VERSION : 0.1
// Data area for auto sequence timers
   VAR
      CV341_CLSD_DLY : TON_TIME;   // For the delay prior to the BC start command
      P305_STRTD_DLY : TON_TIME;   // For the delay after P305 has started
      P304_STRTD_DLY : TON_TIME;   // For the delay after P304 has started
      P303_STRTD_DLY : TON_TIME;   // For the delay after P304 has started
      PRE_GCU_TNK_FILL_DLY : TON_TIME;   // For the delay prior to GCU tank fill timer
      GCU_TNK_MAX_FILL_TMR : TON_TIME;   // For the maximum GCU fill time
      P305_STPD_DLY : TON_TIME;   // For the delay after P305 has stopped
      P304_STPD_DLY : TON_TIME;   // For the delay after P304 has stopped
      CV358_CLSD_DLY : TON_TIME;   // For the delay prior to the BC start command
      E400_STRTD_DLY : TON_TIME;   // For the delay after E400 has started
      E400_RNG_DLY : TON_TIME;   // For the delay as E400 runs at load
      CV401_OPND_DLY : TON_TIME;   // For the delay after CV401 has opened
      CV401_CLSD_DLY : TON_TIME;   // For the delay after CV401 has closed
      CV441_OPND_DLY : TON_TIME;   // For the delay after CV441 has opened
      CV441_CLSD_DLY : TON_TIME;   // For the delay after CV441 has closed
      PRE_441_OPN_DLY : TON_TIME;   // For the delay prior to CV441 opening
      VLV_CNFG_DN_DLY : TON_TIME;   // For the delay once the DeOx/ReOx are done
      CV405_OPND_DLY : TON_TIME;   // For the delay after CV405 has opened
      CV406_CLSD_DLY : TON_TIME;   // For the delay after CV406 has closed
      E400_STOP_TMR : TON_TIME;   // For the maximum PGC stop time
      P303_STPD_DLY : TON_TIME;   // For the maximum P303 stop time
      CV341_OPND_DLY : TON_TIME;   // For the delay after CV341 has opened
      GCU_TNK_MAX_DRN_TMR : TON_TIME;   // For the maximum GCU drain time
      POST_FLUSH_DLY : TON_TIME;   // Dor the delay after the tank has flushed
      "LIT304 Delay" : TON_TIME;
      P301_START_DLY : TON_TIME;   // Delay after starting the CSW pump
      "FS332 Delay" : TON_TIME;
      "Pre-Dwel PPPuls" : TP_TIME;
      SFTY_SYS_IL : TOF_TIME;
      OVR_TANK : TON_TIME;
      "Tank Close Delay" : TON_TIME;
   END_VAR
BEGIN
   CV341_CLSD_DLY.PT := T#10s;
   P305_STRTD_DLY.PT := T#5s;
   P304_STRTD_DLY.PT := T#5s;
   PRE_GCU_TNK_FILL_DLY.PT := T#15s;
   GCU_TNK_MAX_FILL_TMR.PT := T#300s;
   P305_STPD_DLY.PT := T#5s;
   P304_STPD_DLY.PT := T#5s;
   CV358_CLSD_DLY.PT := T#5s;
   P303_STRTD_DLY.PT := T#15s;
   E400_STRTD_DLY.PT := T#15s;
   E400_RNG_DLY.PT := T#5s;
   VLV_CNFG_DN_DLY.PT := T#10s;
   PRE_441_OPN_DLY.PT := T#15s;
   CV441_CLSD_DLY.PT := T#5s;
   CV441_OPND_DLY.PT := T#5s;
   CV401_CLSD_DLY.PT := T#5s;
   CV401_OPND_DLY.PT := T#5s;
   CV405_OPND_DLY.PT := T#10s;
   CV406_CLSD_DLY.PT := T#2s;
   E400_STOP_TMR.PT := T#180s;
   P303_STPD_DLY.PT := T#30s;
   CV341_OPND_DLY.PT := T#2s;
   GCU_TNK_MAX_DRN_TMR.PT := T#180s;
   POST_FLUSH_DLY.PT := T#60s;
   OVR_TANK.PT := T#1s;
   "Tank Close Delay".PT := T#1s;
END_DATA_BLOCK

// folder: 50 - 59 PLC Communication

DATA_BLOCK "51_SLAVE_STATUS"   // DB51
TITLE = Slave Status Data
{ S7_Optimized_Access := 'FALSE' }
AUTHOR : JRS
VERSION : 0.1
// Data area for status from slave PLC
   VAR
      HEART_BEAT : Bool;
      AUT_SEQ_RNG : Bool;   // Auto sequence running
      CRNT_MODE : Int := 1;   // 1 = Auto, 2 = Man, 3 = FatAuto, 4 = FatMan
      STARTING : Bool;   // IGG Is starting
      O2_LVL_OK : Bool;   // O2 Level within specification
      RUNNING : Bool;   // Running
      VLVS_AT_INIT : Bool;   // 1 = Valves at initial, 0 = Not
      ESTOP_OK : Bool;   // 1 = OK, 0 = Estop active
      IGG_ALARM : Bool;   // 1 = IGG Alarm state, 0 = Not
      P305_ENBLD : Bool;   // P305 enabled input sent from BC
      P305_TRIPPED : Bool;   // P305 tripped input sent from BC
      CV401_OPN : Bool;   // CV401 Open
      CV401_CLSD : Bool;   // CV401 Closed
      P301_ENBLD : Bool;   // P305 enabled input sent from BC
      CV311_OPN : Bool;   // CV311 Open
      CV311_CLSD : Bool;   // CV311 CLosed
      CV322_OPN : Bool;   // CV322 Open
      CV322_CLSD : Bool;   // CV322 Closed
      Reset_Alarms : Bool;   // Reset_Alarms
      P305_PRSNT : Bool;   // P305 Present
      ALARM_PRSNT : Bool;   // Alarms from other PLCs
      "CV403 Less 50%" : Bool;
      "BWT Mode Selected" : Bool;
      "CB Mode Selected" : Bool;
      "CV-321_CLSD" : Bool;
      "CAB Started" : Bool;
      "CV403 Opening" : Real;
      "CV431 Opened" : Bool;
      "IGG Stoped" : Bool;
   END_VAR
BEGIN
END_DATA_BLOCK

DATA_BLOCK "56_SLAVE_CMNDS"   // DB56
TITLE = Slave Command Data
{ S7_Optimized_Access := 'FALSE' }
AUTHOR : JRS
VERSION : 0.1
// Data area for commands to slave PLC
   VAR
      HEART_BEAT : Bool;
      CRNT_MODE : Int := 1;   // 1 = Auto, 2 = Man, 3 = FatAuto, 4 = FatMan
      RST_AUT_SEQ : Bool;   // Reset automatic sequence
      GCU_BWT_ALARM : Bool;   // 1 = Alarm, 0 = Not
      OK_RUN_IGG : Bool;   // 1 = Run IGG, 0 = Not
      STOP_IGG : Bool;   // 1 = Stop IGG, 0 = Not
      OPEN_CV401 : Bool;   // 1 = Open, 0 = Not
      RUN_P305 : Bool;   // 1 = Run pump, 0 = Not
      GCU_WRNG_ACTV : Bool;   // 1 = GCU Warning active, 0 = Not
      SPR_BOOL : Bool;   // Spare bit
      RUN_P301 : Bool;   // 1 = Run pump, 0 = Not
      OPEN_CV311 : Bool;   // 1 = Open, 0 = Not
      OPEN_CV322 : Bool;   // 1 = Open, 0 = Not
      NewALARM : Bool;   // NewALARM
      NewWARNING : Bool;   // NewWARNING
      "E-Stop BWT" : Bool;   // E-Stop BWT
      "Mask Interlocks" : Bool;   // Mask Valve Lineup Interlocks for IGG when GCU Shutting Down
      "CV403 Open" : Bool;   // Ctrl from PGC purge FB
      "CV403 Modulate Cmnd" : Bool;   // Ctrl from PGC purge FB
      "CV431 Open Cmd" : Bool;   // Ctrl from PGC purge FB
      "CAB Start Cmd" : Bool;   // Ctrl from PGC purge FB
      "CAB RPM Cmd" : Real;   // Ctrl from PGC purge FB
      "CV401 Open Cmd" : Bool;   // Ctrl from PGC purge FB
   END_VAR
BEGIN
END_DATA_BLOCK

DATA_BLOCK "57_COMMS_DATE_TIME"   // DB57
{ S7_Optimized_Access := 'FALSE' }
VERSION : 0.1
   VAR
      SYSTEM_TIME : DTL;
      LOCAL_TIME : DTL;
   END_VAR
BEGIN
END_DATA_BLOCK

DATA_BLOCK "58_INTRNL_COMMS"   // DB58
TITLE = Internal Communication Data
{ S7_Optimized_Access := 'FALSE' }
AUTHOR : JRS
VERSION : 0.1
// Data area for communication between the BWT and GCU systems within the local PLC
   VAR
      BWT_TO_GCU : Struct
         STATE : Int := 1;   // Current state of BWT
         PREP_GAS : Bool;   // 1 = Prepare gas, 0 = Not
         SPLY_GAS : Bool;   // 1 = Supply gas, 0 = Not
         STP_GAS : Bool;   // 1 = Stop gas, 0 = Not
         FLT_ACTV : Bool;   // 1 = BWT Fault active, 0 = Not
         SHT_DN : Bool;   // 1 = Shutdown, 0 = Not
         SPR_BIT_5 : Bool;   // Spare
         SPR_BIT_6 : Bool;   // Spare
         SPR_BIT_7 : Bool;   // Spare
      END_STRUCT;
      GCU_TO_BWT : Struct
         CRNT_MODE : Int := 1;   // 1 = Auto, 2 = Man, 3 = FatAuto, 4 = FatMan
         PRPNG_GAS : Bool;   // 1 = Preparing gas, 0 = Not
         GAS_AVLBL : Bool;   // 1 = Gas available, 0 = Not
         GAS_DLVRY_ACTV : Bool;   // 1 = Gas delivery active, 0 = Not
         GAS_NOK : Bool;   // 1 = Gas out of specification, 0 = Not
         FLT_ACTV : Bool;   // 1 = BWT Fault active, 0 = Not
         SHT_DN : Bool;   // 1 = Shutdown, 0 = Not
         SPR_BIT_6 : Bool;   // Spare
         SPR_BIT_7 : Bool;   // Spare
      END_STRUCT;
   END_VAR
BEGIN
END_DATA_BLOCK

DATA_BLOCK "59_COMMS_HEALTH_DATA"   // DB59
TITLE = Communications Health Data
{ S7_Optimized_Access := 'TRUE' }
AUTHOR : JRS
VERSION : 0.1
// Data area for communications health determination
   VAR
      CLOCK_POS_EDGE : Bool;
      CLOCK_NEG_EDGE : Bool;
      SLAVE_TRUE_TMR : TON_TIME;
      SLAVE_FALSE_TMR : TON_TIME;
      SLAVE_HB_MISSING : Bool;   // Heartbeat missing flag
   END_VAR
BEGIN
END_DATA_BLOCK

// folder: 60 - 69 Alarm & Satus Handling

DATA_BLOCK "60_Alarm_Data"   // DB60
{ S7_Optimized_Access := 'FALSE' }
VERSION : 0.1
   VAR
      GCU_ALARM_WORD_01 : Word;
      GCU_ALARM_WORD_02 : Word;
      GCU_ALARM_WORD_03 : Word;
      GCU_ALARM_WORD_04 : Word;
      GCU_ALARM_WORD_05 : Word;
      GCU_ALARM_WORD_06 : Word;
      GCU_ALARM_WORD_07 : Word;
      GCU_ALARM_WORD_08 : Word;
      GCU_ALARM_WORD_09 : Word;
      BWTS_ALARM_WORD_10 : Word;
      BWTS_ALARM_WORD_11 : Word;
      BWTS_ALARM_WORD_12 : Word;
      BWTS_ALARM_WORD_13 : Word;
      BWTS_ALARM_WORD_14 : Word;
      BWTS_ALARM_WORD_15 : Word;
      BWTS_ALARM_WORD_16 : Word;
      BWTS_ALARM_WORD_17 : Word;
      BWTS_ALARM_WORD_18 : Word;
      BWTS_ALARM_WORD_19 : Word;
      BWTS_ALARM_WORD_20 : Word;
      BWTS_ALARM_WORD_21 : Word;
      BWTS_ALARM_WORD_22 : Word;
      BWTS_ALARM_WORD_23 : Word;
      BWTS_ALARM_WORD_24 : Word;
      BWTS_ALARM_WORD_25 : Word;
      BWTS_ALARM_WORD_26 : Word;
      BWTS_ALARM_WORD_27 : Word;
      BWTS_ALARM_WORD_28 : Word;
      ALRM_PRSNT : Bool;
      GCU_ALRM_PRSNT : Bool;
      BWTS_ALRM_PRSNT : Bool;
   END_VAR
BEGIN
END_DATA_BLOCK

DATA_BLOCK "Tanks Closed_DB"   // DB61
{ S7_Optimized_Access := 'TRUE' }
VERSION : 0.1
// stored: InstanceOfName Tanks Closed
"Tanks Closed"
BEGIN
END_DATA_BLOCK

DATA_BLOCK "62_Warning_Data"   // DB62
{ S7_Optimized_Access := 'FALSE' }
VERSION : 0.1
   VAR
      GCU_WARNING_WORD_01 : Word;
      GCU_WARNING_WORD_02 : Word;
      GCU_WARNING_WORD_03 : Word;
      GCU_WARNING_WORD_04 : Word;
      GCU_WARNING_WORD_05 : Word;
      GCU_WARNING_WORD_06 : Word;
      GCU_WARNING_WORD_07 : Word;
      GCU_WARNING_WORD_08 : Word;
      GCU_WARNING_WORD_09 : Word;
      BWTS_WARNING_WORD_10 : Word;
      BWTS_WARNING_WORD_11 : Word;
      BWTS_WARNING_WORD_12 : Word;
      BWTS_WARNING_WORD_13 : Word;
      BWTS_WARNING_WORD_14 : Word;
      BWTS_WARNING_WORD_15 : Word;
      BWTS_WARNING_WORD_16 : Word;
      WRNG_PRSNT : Bool;
      GCU_WRNG_PRSNT : Bool;
      BWTS_WRNG_PRSNT : Bool;
   END_VAR
BEGIN
END_DATA_BLOCK

DATA_BLOCK "502_ALM_ANALOG_IDB PIT 353"   // DB63
{ S7_Optimized_Access := 'FALSE' }
VERSION : 0.1
// stored: InstanceOfName 502_ALM_ANALOG
"502_ALM_ANALOG"
BEGIN
END_DATA_BLOCK

DATA_BLOCK "64_Message_Data"   // DB64
{ S7_Optimized_Access := 'FALSE' }
VERSION : 0.1
   VAR
      BWT_MESSAGE_WORD_01 : Word;
      BWT_MESSAGE_WORD_02 : Word;
      BWT_MESSAGE_WORD_03 : Word;
      BWT_MESSAGE_WORD_04 : Word;
      BWT_MESSAGE_WORD_05 : Word;
      BWT_MESSAGE_WORD_06 : Word;
      BWT_MESSAGE_WORD_07 : Word;
      BWT_MESSAGE_WORD_08 : Word;
      MSG_PRSNT : Bool;
   END_VAR
BEGIN
END_DATA_BLOCK

DATA_BLOCK "502_ALM_ANALOG_IDB PIT 416"   // DB65
{ S7_Optimized_Access := 'FALSE' }
VERSION : 0.1
// stored: InstanceOfName 502_ALM_ANALOG
"502_ALM_ANALOG"
BEGIN
END_DATA_BLOCK

DATA_BLOCK "66_Event_Data"   // DB66
{ S7_Optimized_Access := 'FALSE' }
VERSION : 0.1
   VAR
      GCU_EVENT_WORD_01 : Word;
      GCU_EVENT_WORD_02 : Word;
      GCU_EVENT_WORD_03 : Word;
      GCU_EVENT_WORD_04 : Word;
      GCU_EVENT_WORD_05 : Word;
      GCU_EVENT_WORD_06 : Word;
      GCU_EVENT_WORD_07 : Word;
      GCU_EVENT_WORD_08 : Word;
      EVENT_PRSNT : Bool;
   END_VAR
BEGIN
END_DATA_BLOCK

DATA_BLOCK "503_ALARM CHCK_DB"   // DB67
{ S7_Optimized_Access := 'TRUE' }
VERSION : 0.1
// stored: InstanceOfName 503_ALARM CHCK
"503_ALARM CHCK"
BEGIN
END_DATA_BLOCK

DATA_BLOCK "68_Sys_Status_Data"   // DB68
TITLE = System Status Data
{ S7_Optimized_Access := 'TRUE' }
AUTHOR : JRS
VERSION : 0.1
// Data area for system status information as required by the code
   VAR
      VLVS_AT_INIT : Bool;   // All valves at initial position
      INTRLKS_OK : Bool;   // System interlocks ok
      "LOG GCU" : Bool;   // Tag to activate GCU signals logging
      "STOP LOG GCU" : Bool;
      "LOG GCU Simulator" : Bool;
      "NR TANKS ACTIVATED" : Int;
      "NR TANKS ACTIVATED_M" : Int;
      "PIT416_TRGT_RMP_TIME D_INT" : DInt;
      "Tanks Closed" : Bool;
      "Gas to Deck Open" : Bool;
   END_VAR
BEGIN
END_DATA_BLOCK

DATA_BLOCK "503_WARNING CHCK_DB"   // DB69
{ S7_Optimized_Access := 'TRUE' }
VERSION : 0.1
// stored: InstanceOfName 503_ALARM CHCK
"503_ALARM CHCK"
BEGIN
END_DATA_BLOCK

DATA_BLOCK "LIT304_ALM_ANALOG_DB71"   // DB71
{ S7_Optimized_Access := 'FALSE' }
VERSION : 0.1
// stored: InstanceOfName 502_ALM_ANALOG
"502_ALM_ANALOG"
BEGIN
END_DATA_BLOCK

DATA_BLOCK "PIT353_ALM_ANALOG_DB72"   // DB72
{ S7_Optimized_Access := 'FALSE' }
VERSION : 0.1
// stored: InstanceOfName 502_ALM_ANALOG
"502_ALM_ANALOG"
BEGIN
END_DATA_BLOCK

DATA_BLOCK "PIT348_ALM_ANALOG_DB73"   // DB73
{ S7_Optimized_Access := 'FALSE' }
VERSION : 0.1
// stored: InstanceOfName 502_ALM_ANALOG
"502_ALM_ANALOG"
BEGIN
END_DATA_BLOCK

DATA_BLOCK "TIT406_ALM_ANALOG_DB74"   // DB74
{ S7_Optimized_Access := 'FALSE' }
VERSION : 0.1
// stored: InstanceOfName 502_ALM_ANALOG
"502_ALM_ANALOG"
BEGIN
END_DATA_BLOCK

DATA_BLOCK "TIT408_ALM_ANALOG_DB75"   // DB75
{ S7_Optimized_Access := 'FALSE' }
VERSION : 0.1
// stored: InstanceOfName 502_ALM_ANALOG
"502_ALM_ANALOG"
BEGIN
END_DATA_BLOCK

DATA_BLOCK "TT002_ALM_ANALOG_DB76"   // DB76
{ S7_Optimized_Access := 'FALSE' }
VERSION : 0.1
// stored: InstanceOfName 502_ALM_ANALOG
"502_ALM_ANALOG"
BEGIN
END_DATA_BLOCK

DATA_BLOCK "PT002_ALM_ANALOG_DB77"   // DB77
{ S7_Optimized_Access := 'FALSE' }
VERSION : 0.1
// stored: InstanceOfName 502_ALM_ANALOG
"502_ALM_ANALOG"
BEGIN
END_DATA_BLOCK

DATA_BLOCK "PIT358_ALM_ANALOG_DB78"   // DB78
{ S7_Optimized_Access := 'FALSE' }
VERSION : 0.1
// stored: InstanceOfName 502_ALM_ANALOG
"502_ALM_ANALOG"
BEGIN
END_DATA_BLOCK

DATA_BLOCK "HMI Indication Logic_DB"   // DB79
{ S7_Optimized_Access := 'TRUE' }
VERSION : 0.1
// stored: InstanceOfName HMI Indication Logic
"HMI Indication Logic"
BEGIN
END_DATA_BLOCK

DATA_BLOCK "E-400 Animation_DB"   // DB81
{ S7_Optimized_Access := 'TRUE' }
VERSION : 0.1
// stored: InstanceOfName Animation
"Animation"
BEGIN
END_DATA_BLOCK

DATA_BLOCK "FS350 Animation_iDB"   // DB83
{ S7_Optimized_Access := 'TRUE' }
VERSION : 0.1
// stored: InstanceOfName Animation
"Animation"
BEGIN
END_DATA_BLOCK

DATA_BLOCK "FS332 Animation_IDB"   // DB85
{ S7_Optimized_Access := 'TRUE' }
VERSION : 0.1
// stored: InstanceOfName Animation
"Animation"
BEGIN
END_DATA_BLOCK

DATA_BLOCK "P304 Animation_IDB"   // DB87
{ S7_Optimized_Access := 'TRUE' }
VERSION : 0.1
// stored: InstanceOfName Animation
"Animation"
BEGIN
END_DATA_BLOCK

// folder: 70 - 79 Modes of Operation

DATA_BLOCK "70_Mode_Data"   // DB70
{ S7_Optimized_Access := 'TRUE' }
VERSION : 0.1
   VAR
      CRNT_MODE : Int := 1;   // 1 = Auto, 2 = Man, 3 = FatAuto, 4 = FatMan
      INTO_AUTO : Bool;   // Transition to auto
      IN_MAN : Bool;   // In manual
      INTO_AUT_PLS : Bool;   // Pulse bit
      AUT_RST_PLS : TP_TIME;   // Automatic sequence reset pulse
   END_VAR
BEGIN
   AUT_RST_PLS.PT := T#1s;
END_DATA_BLOCK

// folder: 700 - 999 FB Instance DBs

DATA_BLOCK "700_VLV_CHK_DB"   // DB700
{ S7_Optimized_Access := 'TRUE' }
AUTHOR : JRS
VERSION : 0.1
// stored: InstanceOfName 501_VLV_CHK
"501_VLV_CHK"
BEGIN
END_DATA_BLOCK

DATA_BLOCK "701_VLV_CHK_DB"   // DB701
{ S7_Optimized_Access := 'TRUE' }
AUTHOR : JRS
VERSION : 0.1
// stored: InstanceOfName 501_VLV_CHK
"501_VLV_CHK"
BEGIN
END_DATA_BLOCK

DATA_BLOCK "702_VLV_CHK_DB"   // DB702
{ S7_Optimized_Access := 'TRUE' }
AUTHOR : JRS
VERSION : 0.1
// stored: InstanceOfName 501_VLV_CHK
"501_VLV_CHK"
BEGIN
END_DATA_BLOCK

DATA_BLOCK "703_VLV_CHK_DB"   // DB703
{ S7_Optimized_Access := 'TRUE' }
AUTHOR : JRS
VERSION : 0.1
// stored: InstanceOfName 501_VLV_CHK
"501_VLV_CHK"
BEGIN
END_DATA_BLOCK

DATA_BLOCK "704_VLV_CHK_DB"   // DB704
{ S7_Optimized_Access := 'TRUE' }
AUTHOR : JRS
VERSION : 0.1
// stored: InstanceOfName 501_VLV_CHK
"501_VLV_CHK"
BEGIN
END_DATA_BLOCK

DATA_BLOCK "705_VLV_CHK_DB"   // DB705
{ S7_Optimized_Access := 'TRUE' }
AUTHOR : JRS
VERSION : 0.1
// stored: InstanceOfName 501_VLV_CHK
"501_VLV_CHK"
BEGIN
END_DATA_BLOCK

DATA_BLOCK "706_VLV_CHK_DB"   // DB706
{ S7_Optimized_Access := 'TRUE' }
AUTHOR : JRS
VERSION : 0.1
// stored: InstanceOfName 501_VLV_CHK
"501_VLV_CHK"
BEGIN
END_DATA_BLOCK

DATA_BLOCK "720_VLV_CHK_DB"   // DB720
{ S7_Optimized_Access := 'TRUE' }
AUTHOR : JRS
VERSION : 0.1
// stored: InstanceOfName 501_VLV_CHK
"501_VLV_CHK"
BEGIN
END_DATA_BLOCK

// folder: 80 - 89 HMI Handling

DATA_BLOCK "PGC_COMMISSION_MODE_DB"   // DB1
{ S7_Optimized_Access := 'TRUE' }
VERSION : 0.1
   VAR
      Active : Bool;   // Selected from HMI
      Setpoint : Real;   // Commissioning Setpoint from HMI
      "Previous Setpoint" : Real;   // Previous Setpoint from HMI
      "Drive Popup" : Bool;   // Drive Popup to HMI
      "Change SP Pulse" : Bool;   // Pulse to change Setpoint to Commissioning
      "Change SP Back Pulse" : Bool;   // Pulse to change Setpoint to Normal
      "PV Lo Lim" : Real;   // Lower Limit for PV meeting Setpoint
      "PV Hi Lim" : Real;   // Upper Limit for PV meeting Setpoint
      "Button Control" : Int;   // Integer for Button Control
   END_VAR
BEGIN
END_DATA_BLOCK

DATA_BLOCK "PGC_COMMISSION_MODE_TIMER"   // DB2
{ S7_Optimized_Access := 'TRUE' }
AUTHOR : Simatic
FAMILY : IEC
NAME : IEC_TMR
VERSION : 1.0
// stored: InstanceOfName IEC_TIMER
"IEC_TIMER"
BEGIN
END_DATA_BLOCK

DATA_BLOCK "80_From_HMI"   // DB80
TITLE = Data From HMI
{ S7_Optimized_Access := 'TRUE' }
AUTHOR : JRS
VERSION : 0.1
// Data area for signals from the HMI
   VAR
      Request_Manual : Bool := False;   // Pulse from HMI
      Request_Auto : Bool := False;   // Pulse from HMI
      SLNCE_BZR : Bool;   // Pulse to silence buzzer
   END_VAR
   VAR RETAIN
      RUN_BWTS : Bool := false;   // 1 = Run Ballast Water Treatment System, 0 = Not
      RUN_BTCS : Bool := true;   // 1 = Run Barge Tank Control System, 0 = Not
   END_VAR
   VAR
      RST_AUT_SEQ : Bool;   // Reset automatic sequence
      CRG_BLNK_MODE : Bool;   // 1 = Cargon blanketing mode, 0 = Not
   END_VAR
   VAR RETAIN
      P305_PRSNT : Bool := FALSE;   // 1 = Pump fitted, 0 = Not
   END_VAR
   VAR
      STOP_GCU : Bool;   // 1 = Stop, 0 = Not
      SAL_VALUE : Real := 6.0;   // Value to be confirmed
      SAL_CNFRM : Bool;   // Salinity confirmation bit
      LOW_SAL_ACPT : Bool;   // Confirm low salinity
      LOW_SAL_RJCT : Bool;   // Reject low salinity
      PGC_RST_HRS : Bool;   // 1 = Reset Hours, 0 = Not
      P303_RST_HRS : Bool;   // 1 = Reset Hours, 0 = Not
      P304_RST_HRS : Bool;   // 1 = Reset Hours, 0 = Not
      MAN_DQ_136_0 : Bool;   // Q136.0 - Fresh Water Fill Valve Control(CV358)
      MAN_DQ_136_1 : Bool;   // Q136.1 - Waste Water Drain Valve Control (CV341)
      MAN_DQ_136_2 : Bool;   // Q136.2 - Block Valve 1 Control (CV407)
      MAN_DQ_136_3 : Bool;   // Q136.3 - Bleed Valve Control (CV409)
      MAN_DQ_136_4 : Bool;   // Q136.4 - Block Valve 2 Control (CV411)
      MAN_DQ_136_5 : Bool;   // Q136.5 - Ambient Air Valve Control (CV441)
      MAN_DQ_136_6 : Bool;   // Q136.6 - Main Gas to Deck Valve Control (CV406)
      MAN_DQ_136_7 : Bool;   // Q136.7 - Start Process Gas Compressor (E400)
      MAN_DQ_137_0 : Bool;   // Q137.0 - GCU Recirculation Pump Control (P303)
      MAN_DQ_137_1 : Bool;   // Q137.1 - GCU Booster Pump Control (P304)
      MAN_DQ_137_2 : Bool;   // Q137.2 - GCU Warning Alarm (13P1)
      MAN_DQ_137_3 : Bool;   // Q137.3 - GCU Shutdown Alarm (13P2)
      MAN_DQ_137_4 : Bool;   // Q137.4 - GCU Running (13P3)
      MAN_DQ_137_5 : Bool;   // Q137.5 - Ballast Water Tank Level High High (13P4)
      MAN_DQ_137_6 : Bool;   // Q137.6 - GCU Alarm Buzzer (13P5)
      MAN_DQ_137_7 : Bool;   // Q137.7 - Stop Process Gas Compressor (E400)
      MAN_DQ_138_0 : Bool;   // Q138.0 - Pilot For GTT FPT Valve (CV422-FPT)
      MAN_DQ_138_1 : Bool;   // Q138.1 - Pilot For GTT 1 Port Valve (CV422-1P)
      MAN_DQ_138_2 : Bool;   // Q138.2 - Pilot For GTT 1 Starboard Valve (CV421-1S)
      MAN_DQ_138_3 : Bool;   // Q138.3 - Pilot For GTT 2 Port Valve (CV422-2P)
      MAN_DQ_138_4 : Bool;   // Q138.4 - Pilot For GTT 2 Starboard Valve (CV421-2S)
      MAN_DQ_138_5 : Bool;   // Q138.5 - Pilot For GTT 3 Port Valve (CV422-3P)
      MAN_DQ_138_6 : Bool;   // Q138.6 - Pilot For GTT 3 Starboard Valve (CV421-3S)
      MAN_DQ_138_7 : Bool;   // Q138.7 - Spare Output
      MAN_DQ_139_0 : Bool;   // Q139.0 - Pilot For GTT 4 Port Valve (CV422-4P)
      MAN_DQ_139_1 : Bool;   // Q139.1 - Pilot For GTT 4 Starboard Valve (CV421-4S)
      MAN_DQ_139_2 : Bool;   // Q139.2 - Pilot For GTT 5 Port Valve (CV422-5P)
      MAN_DQ_139_3 : Bool;   // Q139.3 - Pilot For GTT 5 Starboard Valve (CV421-5S)
      MAN_DQ_139_4 : Bool;   // Q139.4 - Pilot For GTT 6 Port Valve (CV422-6P)
      MAN_DQ_139_5 : Bool;   // Q139.5 - Pilot For GTT 6 Starboard Valve (CV421-6S)
      MAN_DQ_139_6 : Bool;   // Q139.6 - Pilot For GTT APT Valve (CV422-APT)
      MAN_DQ_139_7 : Bool;   // Q139.7 - Spare Output
      MAN_AQ_INC_800 : Bool;   // QW800 - CV405 - Increase % Signal
      MAN_AQ_DEC_800 : Bool;   // QW800 - CV405 - Decrease % Signal
      MAN_AQ_INC_802 : Bool;   // QW802 - Spare - Increase % Signal
      MAN_AQ_DEC_802 : Bool;   // QW802 - Spare - Decrease % Signal
      MAN_AQ_INC_804 : Bool;   // QW804 - Spare - Increase % Signal
      MAN_AQ_DEC_804 : Bool;   // QW804 - Spare - Decrease % Signal
      MAN_AQ_INC_806 : Bool;   // QW806 - Spare - Increase % Signal
      MAN_AQ_DEC_806 : Bool;   // QW806 - Spare - Decrease % Signal
      "TIMER RST Supres" : Bool;
      "Test Tank Request" : Bool;
   END_VAR
   VAR RETAIN
      "m³/hr to Nm³/hr" : Bool := FALSE;
   END_VAR
   VAR
      "Jurney Start Simulator" : Bool;
   END_VAR
   VAR RETAIN
      "TT002 Target Protection" : Bool := TRUE;   // Activate PGC Temperature Protection
      "PT002 Target Protection" : Bool := TRUE;   // Activate PGC Presure Protection
      "Tank Close Protection" : Bool := TRUE;   // Activate Tank Change Pressure Setpoint protection
   END_VAR
   VAR
      "GCU Start Confirmed" : Bool;
   END_VAR
BEGIN
END_DATA_BLOCK

DATA_BLOCK "82_To_HMI"   // DB82
TITLE = Data To HMI
{ S7_Optimized_Access := 'TRUE' }
AUTHOR : JRS
VERSION : 0.1
// Data area for signals to the HMI
   VAR
      CRNT_MODE_GCU : Int := 1;   // 1 = Man, 2 = Auto, 3 = FAT Man, 4 = FATAuto
      AUTO_SEQ_RNG : Bool;   // 1 = Auto sequence running, 0 = Not
      "FS350 Animation" : Int;
      "FS332 Animation" : Int;
      "P304 Animation" : Int;
      "Re-Ox Warning" : Bool;
      "Warn to Start IGG" : Bool;
      "Warn to Start IGG-Last" : Bool;
      "Warn to Start GCU" : Bool;
      "Warn to Start GCU-Last" : Bool;
   END_VAR
BEGIN
END_DATA_BLOCK

DATA_BLOCK "84_Setpoints"   // DB84
TITLE = Setpoints Data
{ S7_Optimized_Access := 'TRUE' }
AUTHOR : JRS
VERSION : 0.1
// Setpoints data area
   VAR RETAIN
      LIT304_InitialFill_Target : Real := 60.0;   // LIT304 initial fill target (%) [GEN-19]
      LIT304_InitialFill_Target_Low : Real := 55.0;
      LIT304_InitialFill_LowLow : Real := 10.0;   // LIT304 initial fill low low setpoint (%) [GEN-19]
      LIT304_InitialFill_Low : Real := 20.0;   // LIT304 initial fill low set point (%) [GEN-19]
      LIT304_InitialFill_High : Real := 80.0;   // LIT304 initial fill high setpoint (%) [GEN-19]
      LIT304_InitialFill_HighHigh : Real := 90.0;   // LIT304 initial fill high high setpoint (%)
      LIT304_Refill_Target : Real := 50.0;   // LIT304 refill target setpoint (%)
      LIT304_Refill_Target_Low : Real := 30.0;
      LIT304_Refill_LowLow : Real := 10.0;   // LIT304 refill low low setpoint (%)
      LIT304_Refill_Low : Real := 20.0;   // LIT304 refill low setpoint (%)
      LIT304_Refill_High : Real := 80.0;   // LIT304 refill high setpoint (%)
      LIT304_Refill_HighHigh : Real := 90.0;   // LIT304 refill high high setpoint (%)
      PIT416_Target : Real := 3.2;   // PIT416 target setpoint (bar g)
      PIT416_LowLow : Real := 0.3;   // PIT416 low low setpoint (bar g)
      PIT416_Low : Real := 0.4;   // PIT416 low setpoint (bar g)
      PIT416_High : Real := 4.5;   // PIT416 high setpoint (bar g)
      PIT416_HighHigh : Real := 4.8;   // PIT416 high high setpoint (bar g)
      TIT406_High : Real := 65.0;   // TIT406 high setpoint (degC)
      TIT406_HighHigh : Real := 70.0;   // TIT406 high high setpoint (degC)
      TIT408_High : Real := 45.0;   // TIT408 high setpoint (degC)
      TIT408_HighHigh : Real := 50.0;   // TIT408 high high setpoint (degC)
      PIT353_InitialFill_LowLow : Real := 0.2;   // PIT353 initial fill low low setpoint (bar g)
      PIT353_InitialFill_Low : Real := 0.3;   // PIT353 initial fill low setpoint (bar g)
      PIT353_InitialFill_High : Real := 6.0;   // PIT353 initial fill high setpoint (bar g)
      PIT353_InitialFill_HighHigh : Real := 6.2;   // PIT353 initial fill high high setpoint (bar g)
      PIT353_Refill_LowLow : Real := 0.2;   // PIT353 refill low low setpoint (bar g)
      PIT353_Refill_Low : Real := 0.4;   // PIT353 refill low setpoint (bar g)
      PIT353_Refill_High : Real := 6.0;   // PIT353 refill high setpoint (bar g)
      PIT353_Refill_HighHigh : Real := 6.2;   // PIT353 refill high high setpoint (bar g)
      PIT348_LowLow : Real := 0.1;   // PIT348 low low setpoint (bar g)
      PIT348_Low : Real := 0.2;   // PIT348 low setpoint (bar g)
      PIT348_High : Real := 2.5;   // PIT348 high setpoint (bar g)
      PIT348_HighHigh : Real := 3.0;   // PIT348 high high setpoint (bar g)
      PIT358_InitialFill_LowLow : Real := 0.2;   // PIT358 initial fill low low setpoint (bar g)
      PIT358_InitialFill_Low : Real := 0.3;   // PIT358 initial fill low setpoint (bar g)
      PIT358_InitialFill_High : Real := 10.0;   // PIT358 initial fill high setpoint (bar g)
      PIT358_InitialFill_HighHigh : Real := 11.0;   // PIT358 initial fill high high setpoint (bar g)
      PIT358_Refill_LowLow : Real := 0.7;   // PIT358 refill low low setpoint (bar g)
      PIT358_Refill_Low : Real := 0.8;   // PIT358 refill low setpoint (bar g)
      PIT358_Refill_High : Real := 10.0;   // PIT358 refill high setpoint (bar g)
      PIT358_Refill_HighHigh : Real := 11.0;   // PIT358 refill high high setpoint (bar g)
      E400_PT002_High : Real := 4.5;   // PT002 PGC Outlet pressure high setpoint (bar g)
      E400_PT002_HighHigh : Real := 4.8;   // PT002 PGC Outlet pressure highhigh setpoint (bar g)
      E400_TT002_High : Real := 250.0;   // TT002 PGC Outlet temperature high setpoint (deg c)
      E400_TT002_HighHigh : Real := 270.0;   // TT002 PGC Outlet temperature highhigh setpoint (deg c)
      NumberCWPumps : Int := 1;   // Number of CW Pumps
      GCUCWPumpCHM : Bool := FALSE;   // True = CHM supplied pump, False = ship supplied pump
      PIT416_Target_Safe : Real := 2.0;   // PIT416 target safe setpoint (bar g)
      "E-400 TT002 Tolerance" : Real := 10.0;   // PGC Temperature Tolerance
      "E-400 PT002 Tolerance" : Real := 0.1;   // PGC Pressure Tolerance
      "Tank Close TimeOut" : Time := T#1M;   // Tank Change Pressure Setpoint protection Time
   END_VAR
BEGIN
END_DATA_BLOCK

DATA_BLOCK "86_Times"   // DB86
TITLE = Times Data
{ S7_Optimized_Access := 'TRUE' }
AUTHOR : JRS
VERSION : 0.1
// Times data area
   VAR RETAIN
      P303_STRTD_DLY : Time := T#15S;   // Sequence step delay time
      P303_STPD_DLY : Time := T#5S;   // Sequence step delay time
      P304_STRTD_DLY : Time := T#5S;   // Sequence step delay time
      P304_STPD_DLY : Time := T#5S;   // Sequence step delay time
      P305_STRTD_DLY : Time := T#5S;   // Sequence step delay time
      P305_STPD_DLY : Time := T#5S;   // Sequence step delay time
      CV341_CLSD_DLY : Time := T#5S;   // Sequence step delay time
      CV358_CLSD_DLY : Time := T#5S;   // Sequence step delay time
      CV401_OPND_DLY : Time := T#0MS;   // Sequence step delay time
      CV401_CLSD_DLY : Time := T#5S;   // Sequence step delay time
      CV441_OPND_DLY : Time := T#0MS;   // Sequence step delay time
      CV441_CLSD_DLY : Time := T#5S;   // Sequence step delay time
      PRE_CV441_OPN_DLY : Time := T#0MS;   // Sequence step delay time
      VLV_CNFG_DN_DLY : Time := T#10S;   // Sequence step delay time
      PRE_GCU_TNK_FILL_DLY : Time := T#15S;   // Sequence step delay time
      GCU_TNK_FILL_MAX_TIME : Time := T#10M;   // GCU Tank maximum fill time
      E400_STRTD_DLY : Time := T#15S;   // Sequence step delay time
      E400_RNG_DLY : Time := T#1S;   // Sequence step delay time
      CV405_OPND_DLY : Time := T#10S;   // Sequence step delay time
      CV406_CLSD_DLY : Time := T#10S;   // Sequence step delay time
      E400_STOP_TIME : Time := T#3M;   // E400 (PGC) Maximum stop time
      P303_STOP_TIME : Time := T#30S;   // P303 Maximum stop time
      CV341_OPND_DLY : Time := T#10S;   // Sequence step delay time
      GCU_TNK_DRN_MAX_TIME : Time := T#2M;   // GCU Tank maximum drain time
      GCU_FLUSH_TIME : Time := T#30S;   // Flush time
      POST_FLUSH_DLY : Time := T#15S;   // Sequence step delay time
      CV341_MAX_TRVL_TIME : Time := T#30S;   // Maximum valve travel time
      CV358_MAX_TRVL_TIME : Time := T#30S;   // Maximum valve travel time
      CV406_MAX_TRVL_TIME : Time := T#30S;   // Maximum valve travel time
      CV407_MAX_TRVL_TIME : Time := T#30S;   // Maximum valve travel time
      CV409_MAX_TRVL_TIME : Time := T#30S;   // Maximum valve travel time
      CV411_MAX_TRVL_TIME : Time := T#30S;   // Maximum valve travel time
      CV441_MAX_TRVL_TIME : Time := T#30S;   // Maximum valve travel time
      PIT416_TRGT_RMP_TIME : Real := 30.0;   // Target Ramp Time In Seconds
      STEP_MAX_TIME_STP_001 : Time := T#30MS;   // Maximum sequence step time
      STEP_MAX_TIME_STP_005 : Time := T#30MS;   // Maximum sequence step time
      STEP_MAX_TIME_STP_010 : Time := T#30MS;   // Maximum sequence step time
      STEP_MAX_TIME_STP_020 : Time := T#30MS;   // Maximum sequence step time
      STEP_MAX_TIME_STP_030 : Time := T#30MS;   // Maximum sequence step time
      STEP_MAX_TIME_STP_040 : Time := T#30MS;   // Maximum sequence step time
      STEP_MAX_TIME_STP_050 : Time := T#30MS;   // Maximum sequence step time
      STEP_MAX_TIME_STP_060 : Time := T#30MS;   // Maximum sequence step time
      STEP_MAX_TIME_STP_070 : Time := T#30MS;   // Maximum sequence step time
      STEP_MAX_TIME_STP_080 : Time := T#30MS;   // Maximum sequence step time
      STEP_MAX_TIME_STP_090 : Time := T#30MS;   // Maximum sequence step time
      STEP_MAX_TIME_STP_100 : Time := T#30MS;   // Maximum sequence step time
      STEP_MAX_TIME_STP_110 : Time := T#30MS;   // Maximum sequence step time
      STEP_MAX_TIME_STP_120 : Time := T#30MS;   // Maximum sequence step time
      STEP_MAX_TIME_STP_130 : Time := T#30MS;   // Maximum sequence step time
      STEP_MAX_TIME_STP_140 : Time := T#30MS;   // Maximum sequence step time
      STEP_MAX_TIME_STP_150 : Time := T#30MS;   // Maximum sequence step time
      STEP_MAX_TIME_STP_160 : Time := T#30MS;   // Maximum sequence step time
      STEP_MAX_TIME_STP_170 : Time := T#30MS;   // Maximum sequence step time
      STEP_MAX_TIME_STP_180 : Time := T#30MS;   // Maximum sequence step time
      STEP_MAX_TIME_STP_190 : Time := T#30MS;   // Maximum sequence step time
      STEP_MAX_TIME_STP_200 : Time := T#30MS;   // Maximum sequence step time
      STEP_MAX_TIME_STP_210 : Time := T#30MS;   // Maximum sequence step time
      STEP_MAX_TIME_STP_220 : Time := T#30MS;   // Maximum sequence step time
      STEP_MAX_TIME_STP_230 : Time := T#30MS;   // Maximum sequence step time
      STEP_MAX_TIME_STP_240 : Time := T#30MS;   // Maximum sequence step time
      STEP_MAX_TIME_STP_250 : Time := T#30MS;   // Maximum sequence step time
      STEP_MAX_TIME_STP_260 : Time := T#30MS;   // Maximum sequence step time
      STEP_MAX_TIME_STP_270 : Time := T#30MS;   // Maximum sequence step time
      STEP_MAX_TIME_STP_280 : Time := T#30MS;   // Maximum sequence step time
      STEP_MAX_TIME_STP_290 : Time := T#30MS;   // Maximum sequence step time
      STEP_MAX_TIME_STP_300 : Time := T#30MS;   // Maximum sequence step time
      STEP_MAX_TIME_STP_310 : Time := T#30MS;   // Maximum sequence step time
      STEP_MAX_TIME_STP_320 : Time := T#3S;   // Maximum sequence step time
      STEP_MAX_TIME_STP_330 : Time := T#30MS;   // Maximum sequence step time
      STEP_MAX_TIME_STP_340 : Time := T#30MS;   // Maximum sequence step time
      STEP_MAX_TIME_STP_350 : Time := T#30MS;   // Maximum sequence step time
      STEP_MAX_TIME_STP_360 : Time := T#30MS;   // Maximum sequence step time
      STEP_MAX_TIME_STP_370 : Time := T#3S;   // Maximum sequence step time
      STEP_MAX_TIME_STP_380 : Time := T#30MS;   // Maximum sequence step time
      STEP_MAX_TIME_STP_390 : Time := T#30MS;   // Maximum sequence step time
      STEP_MAX_TIME_STP_400 : Time := T#30MS;   // Maximum sequence step time
      STEP_MAX_TIME_STP_410 : Time := T#30MS;   // Maximum sequence step time
      STEP_MAX_TIME_STP_420 : Time := T#30MS;   // Maximum sequence step time
      STEP_MAX_TIME_STP_430 : Time := T#30MS;   // Maximum sequence step time
      STEP_MAX_TIME_STP_440 : Time := T#30MS;   // Maximum sequence step time
      STEP_MAX_TIME_STP_450 : Time := T#30MS;   // Maximum sequence step time
      STEP_MAX_TIME_STP_460 : Time := T#30MS;   // Maximum sequence step time
      STEP_MAX_TIME_STP_470 : Time := T#30MS;   // Maximum sequence step time
      STEP_MAX_TIME_STP_480 : Time := T#30MS;   // Maximum sequence step time
      STEP_MAX_TIME_STP_490 : Time := T#30MS;   // Maximum sequence step time
      STEP_MAX_TIME_STP_500 : Time := T#30MS;   // Maximum sequence step time
      STEP_MAX_TIME_STP_510 : Time := T#3S;   // Maximum sequence step time
      STEP_MAX_TIME_STP_520 : Time := T#30MS;   // Maximum sequence step time
      STEP_MAX_TIME_STP_530 : Time := T#3M;   // Maximum sequence step time
      STEP_MAX_TIME_STP_540 : Time := T#30MS;   // Maximum sequence step time
      STEP_MAX_TIME_STP_550 : Time := T#30MS;   // Maximum sequence step time
      STEP_MAX_TIME_STP_560 : Time := T#30MS;   // Maximum sequence step time
      STEP_MAX_TIME_STP_570 : Time := T#30MS;   // Maximum sequence step time
      STEP_MAX_TIME_STP_580 : Time := T#30MS;   // Maximum sequence step time
      STEP_MAX_TIME_STP_590 : Time := T#30MS;   // Maximum sequence step time
      STEP_MAX_TIME_STP_600 : Time := T#30MS;   // Maximum sequence step time
      STEP_MAX_TIME_STP_610 : Time := T#30MS;   // Maximum sequence step time
      STEP_MAX_TIME_STP_620 : Time := T#30MS;   // Maximum sequence step time
      STEP_MAX_TIME_STP_630 : Time := T#30MS;   // Maximum sequence step time
   END_VAR
   VAR
      "PIT353 Delay" : Time := T#10S;
      "PIT416 Delay" : Time := T#10S;
      P301_START_DLY : Time := T#15S;
      "FS332 Delay" : Time := T#10S;
      "LIT304 Delay" : Time := T#10S;
      "PIT358 Delay" : Time := T#30S;   // Fresh Water Inlet Pressure Alarm Delay
      "PIT348 Delay" : Time := T#10S;   // Cooling Seawater Pressure Alarm Delay
   END_VAR
BEGIN
END_DATA_BLOCK

DATA_BLOCK "88_treatment"   // DB88
{ S7_Optimized_Access := 'TRUE' }
VERSION : 0.1
   VAR
      POP_UP : Bool;
      POP_UP_CNFRM : Bool;
   END_VAR
BEGIN
END_DATA_BLOCK

// folder: 90 - 99 Manual Functions

DATA_BLOCK "90_Manual_Data"   // DB90
{ S7_Optimized_Access := 'TRUE' }
VERSION : 0.1
   VAR
      INC_PLS_800 : Bool;   // Pulse bit
      INC_PLS_800_Hz : Bool;   // Pulse bit
      DEC_PLS_800 : Bool;   // Pulse bit
      DEC_PLS_800_Hz : Bool;   // Pulse bit
      INC_PLS_802 : Bool;   // Pulse bit
      INC_PLS_802_Hz : Bool;   // Pulse bit
      DEC_PLS_802 : Bool;   // Pulse bit
      DEC_PLS_802_Hz : Bool;   // Pulse bit
      INC_PLS_804 : Bool;   // Pulse bit
      INC_PLS_804_Hz : Bool;   // Pulse bit
      DEC_PLS_804 : Bool;   // Pulse bit
      DEC_PLS_804_Hz : Bool;   // Pulse bit
      INC_PLS_806 : Bool;   // Pulse bit
      INC_PLS_806_Hz : Bool;   // Pulse bit
      DEC_PLS_806 : Bool;   // Pulse bit
      DEC_PLS_806_Hz : Bool;   // Pulse bit
   END_VAR
BEGIN
END_DATA_BLOCK

// folder: System blocks/Program resources

DATA_BLOCK "IEC_Timer_0_DB"   // DB3
{ S7_Optimized_Access := 'TRUE' }
AUTHOR : Simatic
FAMILY : IEC
NAME : IEC_TMR
VERSION : 1.0
// stored: InstanceOfName IEC_TIMER
"IEC_TIMER"
BEGIN
END_DATA_BLOCK

DATA_BLOCK "IEC_Timer_0_DB_1"   // DB4
{ S7_Optimized_Access := 'TRUE' }
AUTHOR : Simatic
FAMILY : IEC
NAME : IEC_TMR
VERSION : 1.0
// stored: InstanceOfName IEC_TIMER
"IEC_TIMER"
BEGIN
END_DATA_BLOCK

// folder: (top level)

ORGANIZATION_BLOCK "BWTS Main"   // OB1, LAD, ProgramCycle
TITLE = "Main Program Sweep (Cycle)"
{ S7_Optimized_Access := 'FALSE' }
VERSION : 0.1
   VAR_TEMP
      OB1_EV_CLASS : Byte;   // Bits 0-3 = 1 (Coming event), Bits 4-7 = 1 (Event class 1)
      OB1_SCAN_1 : Byte;   // 1 (Cold restart scan 1 of OB 1), 3 (Scan 2-n of OB 1)
      OB1_PRIORITY : Byte;   // Priority of OB Execution
      OB1_OB_NUMBR : Byte;   // 1 (Organization block 1, OB1)
      OB1_RESERVED_1 : Byte;   // Reserved for system
      OB1_RESERVED_2 : Byte;   // Reserved for system
      OB1_PREV_CYCLE : Int;   // Cycle time of previous OB1 scan (milliseconds)
      OB1_MIN_CYCLE : Int;   // Minimum cycle time of OB1 (milliseconds)
      OB1_MAX_CYCLE : Int;   // Maximum cycle time of OB1 (milliseconds)
      OB1_DATE_TIME : Date_And_Time;   // Date and time OB1 started
   END_VAR
   VAR_TEMP   // added for the SCL form of the ladder/FBD networks
      _w1 : Bool;
   END_VAR
BEGIN

REGION Network 1: Digital Input Processing
   // To process raw inputs prior to code use